   Reference[401].Actionpoint_2[7] := '0';
   Reference[401].Actionpoint_2[6] := '0';
   Reference[401].Actionpoint_2[5] := '0';
   Reference[401].Actionpoint_2[4] := '0';
   Reference[401].Actionpoint_2[3] := '0';
   Reference[401].Actionpoint_2[2] := '0';
   Reference[401].Actionpoint_2[1] := '0';
   Reference[401].Actionpoint_1[16] := '0';
   Reference[401].Actionpoint_1[15] := '0';
   Reference[401].Actionpoint_1[14] := '0';
   Reference[401].Actionpoint_1[13] := '0';
   Reference[401].Actionpoint_1[12] := '0';
   Reference[401].Actionpoint_1[11] := '0';
   Reference[401].Actionpoint_1[10] := '0';
   Reference[401].Actionpoint_1[9] := '0';
   Reference[401].Actionpoint_1[8] := '0';
   Reference[401].Actionpoint_1[7] := '0';
   Reference[401].Actionpoint_1[6] := '0';
   Reference[401].Actionpoint_1[5] := '0';
   Reference[401].Actionpoint_1[4] := '0';
   Reference[401].Actionpoint_1[3] := '0';
   Reference[401].Actionpoint_1[2] := '0';
   Reference[401].Actionpoint_1[1] := '0';
   Reference[401].Sektion[1] := 'b';
   Reference[401].Sektion[2] := 'u';
   Reference[401].Sektion[3] := 'f';
   Reference[401].Sektion[4] := 'f';
   Reference[401].Sektion[5] := 'e';
   Reference[401].Sektion[6] := 'r';
   Reference[401].Sektion[7] := '$00';
   Reference[401].Sektion[8] := '$00';
   Reference[401].Sektion[9] := '$00';
   Reference[401].Sektion[10] := '$00';
   Reference[401].Sektion[11] := '$00';
   Reference[401].Sektion[12] := '$00';
   Reference[401].Sektion[13] := '$00';
   Reference[401].Sektion[14] := '$00';
   Reference[401].Sektion[15] := '$00';
   Reference[401].Sektion[16] := '$00';
   // 19800 more start values not shown
END_DATA_BLOCK

DATA_BLOCK "DB_SDC_TS_REFERENCE_6"   // DB3785
{ S7_Optimized_Access := 'FALSE' }
VERSION : 0.1
   VAR
      HEADER : Struct   // Struktur für Datenheader // nicht verschieben
         DB_NR : Int := 3785;   // DB Nummer
         MIN_NR_SEK : Int := 501;   // Niedrigste SEK Nummer im DB
         MAX_NR_SEK : Int := 600;   // Höchste SEK Nummer im DB
         START_DAT : Int := 20;   // Startadresse der SEK im DB
         LAENGE_SEK_DATA : Int := 200;   // Länge SEK Data
         Res10 : Int := 0;   // Reserve
         Res12 : Int := 0;   // Reserve
         Res14 : Int := 0;   // Reserve
         Res16 : Int := 0;   // Reserve
         Res18 : Int := 0;   // Reserve
      END_STRUCT;
      Reference : Array[501..600] of Struct   // Sektionsnummer
         Sektion : Array[1..16] of Char;   // definition Sektion
         Actionpoint_1 : Array[1..16] of Char;   // definition Actionpoint 1
         Actionpoint_2 : Array[1..16] of Char;   // definition Actionpoint 2
         Height : Array[1..16] of Char;   // definition Hubposition (mm)
         Hoist_offset_1 : Array[1..16] of Char;   // definition Hub-Offset 1 (mm)
         Hoist_offset_2 : Array[1..16] of Char;   // definition Hub-Offset 2 (mm)
         Hoist_offset_3 : Array[1..16] of Char;   // definition Hub-Offset 3(mm)
         Hoist_offset_4 : Array[1..16] of Char;   // definition Hub-Offset 4 (mm)
         Reserve : Array[128..199] of Char;
      END_STRUCT;
   END_VAR
BEGIN
   Reference[501].Reserve[199] := ' ';
   Reference[501].Reserve[198] := ' ';
   Reference[501].Reserve[197] := ' ';
   Reference[501].Reserve[196] := ' ';
   Reference[501].Reserve[195] := ' ';
   Reference[501].Reserve[194] := ' ';
   Reference[501].Reserve[193] := ' ';
   Reference[501].Reserve[192] := ' ';
   Reference[501].Reserve[191] := ' ';
   Reference[501].Reserve[190] := ' ';
   Reference[501].Reserve[189] := ' ';
   Reference[501].Reserve[188] := ' ';
   Reference[501].Reserve[187] := ' ';
   Reference[501].Reserve[186] := ' ';
   Reference[501].Reserve[185] := ' ';
   Reference[501].Reserve[184] := ' ';
   Reference[501].Reserve[183] := ' ';
   Reference[501].Reserve[182] := ' ';
   Reference[501].Reserve[181] := ' ';
   Reference[501].Reserve[180] := ' ';
   Reference[501].Reserve[179] := ' ';
   Reference[501].Reserve[178] := ' ';
   Reference[501].Reserve[177] := ' ';
   Reference[501].Reserve[176] := ' ';
   Reference[501].Reserve[175] := ' ';
   Reference[501].Reserve[174] := ' ';
   Reference[501].Reserve[173] := ' ';
   Reference[501].Reserve[172] := ' ';
   Reference[501].Reserve[171] := ' ';
   Reference[501].Reserve[170] := ' ';
   Reference[501].Reserve[169] := ' ';
   Reference[501].Reserve[168] := ' ';
   Reference[501].Reserve[167] := ' ';
   Reference[501].Reserve[166] := ' ';
   Reference[501].Reserve[165] := ' ';
   Reference[501].Reserve[164] := ' ';
   Reference[501].Reserve[163] := ' ';
   Reference[501].Reserve[162] := ' ';
   Reference[501].Reserve[161] := ' ';
   Reference[501].Reserve[160] := ' ';
   Reference[501].Reserve[159] := ' ';
   Reference[501].Reserve[158] := ' ';
   Reference[501].Reserve[157] := ' ';
   Reference[501].Reserve[156] := ' ';
   Reference[501].Reserve[155] := ' ';
   Reference[501].Reserve[154] := ' ';
   Reference[501].Reserve[153] := ' ';
   Reference[501].Reserve[152] := ' ';
   Reference[501].Reserve[151] := ' ';
   Reference[501].Reserve[150] := ' ';
   Reference[501].Reserve[149] := ' ';
   Reference[501].Reserve[148] := ' ';
   Reference[501].Reserve[147] := ' ';
   Reference[501].Reserve[146] := ' ';
   Reference[501].Reserve[145] := ' ';
   Reference[501].Reserve[144] := ' ';
   Reference[501].Reserve[143] := '0';
   Reference[501].Reserve[142] := '0';
   Reference[501].Reserve[141] := '0';
   Reference[501].Reserve[140] := '0';
   Reference[501].Reserve[139] := '0';
   Reference[501].Reserve[138] := '0';
   Reference[501].Reserve[137] := '0';
   Reference[501].Reserve[136] := '0';
   Reference[501].Reserve[135] := '0';
   Reference[501].Reserve[134] := '0';
   Reference[501].Reserve[133] := '0';
   Reference[501].Reserve[132] := '0';
   Reference[501].Reserve[131] := '0';
   Reference[501].Reserve[130] := '0';
   Reference[501].Reserve[129] := '0';
   Reference[501].Reserve[128] := '0';
   Reference[501].Hoist_offset_4[16] := '$00';
   Reference[501].Hoist_offset_4[15] := '$00';
   Reference[501].Hoist_offset_4[14] := '$00';
   Reference[501].Hoist_offset_4[13] := '$00';
   Reference[501].Hoist_offset_4[12] := '$00';
   Reference[501].Hoist_offset_4[11] := '$00';
   Reference[501].Hoist_offset_4[10] := '$00';
   Reference[501].Hoist_offset_4[9] := '$00';
   Reference[501].Hoist_offset_4[8] := '$00';
   Reference[501].Hoist_offset_4[7] := '$00';
   Reference[501].Hoist_offset_4[6] := '$00';
   Reference[501].Hoist_offset_4[5] := '$00';
   Reference[501].Hoist_offset_4[4] := '$00';
   Reference[501].Hoist_offset_4[3] := '$00';
   Reference[501].Hoist_offset_4[2] := '$00';
   Reference[501].Hoist_offset_4[1] := '$00';
   Reference[501].Hoist_offset_3[16] := '$00';
   Reference[501].Hoist_offset_3[15] := '$00';
   Reference[501].Hoist_offset_3[14] := '$00';
   Reference[501].Hoist_offset_3[13] := '$00';
   Reference[501].Hoist_offset_3[12] := '$00';
   Reference[501].Hoist_offset_3[11] := '$00';
   Reference[501].Hoist_offset_3[10] := '$00';
   Reference[501].Hoist_offset_3[9] := '$00';
   Reference[501].Hoist_offset_3[8] := '$00';
   Reference[501].Hoist_offset_3[7] := '$00';
   Reference[501].Hoist_offset_3[6] := '$00';
   Reference[501].Hoist_offset_3[5] := '$00';
   Reference[501].Hoist_offset_3[4] := '$00';
   Reference[501].Hoist_offset_3[3] := '$00';
   Reference[501].Hoist_offset_3[2] := '$00';
   Reference[501].Hoist_offset_3[1] := '$00';
   Reference[501].Hoist_offset_2[16] := '$00';
   Reference[501].Hoist_offset_2[15] := '$00';
   Reference[501].Hoist_offset_2[14] := '$00';
   Reference[501].Hoist_offset_2[13] := '$00';
   Reference[501].Hoist_offset_2[12] := '$00';
   Reference[501].Hoist_offset_2[11] := '$00';
   Reference[501].Hoist_offset_2[10] := '$00';
   Reference[501].Hoist_offset_2[9] := '$00';
   Reference[501].Hoist_offset_2[8] := '$00';
   Reference[501].Hoist_offset_2[7] := '$00';
   Reference[501].Hoist_offset_2[6] := '$00';
   Reference[501].Hoist_offset_2[5] := '$00';
   Reference[501].Hoist_offset_2[4] := '$00';
   Reference[501].Hoist_offset_2[3] := '$00';
   Reference[501].Hoist_offset_2[2] := '$00';
   Reference[501].Hoist_offset_2[1] := '$00';
   Reference[501].Hoist_offset_1[16] := '$00';
   Reference[501].Hoist_offset_1[15] := '$00';
   Reference[501].Hoist_offset_1[14] := '$00';
   Reference[501].Hoist_offset_1[13] := '$00';
   Reference[501].Hoist_offset_1[12] := '$00';
   Reference[501].Hoist_offset_1[11] := '$00';
   Reference[501].Hoist_offset_1[10] := '$00';
   Reference[501].Hoist_offset_1[9] := '$00';
   Reference[501].Hoist_offset_1[8] := '$00';
   Reference[501].Hoist_offset_1[7] := '$00';
   Reference[501].Hoist_offset_1[6] := '$00';
   Reference[501].Hoist_offset_1[5] := '$00';
   Reference[501].Hoist_offset_1[4] := '$00';
   Reference[501].Hoist_offset_1[3] := '$00';
   Reference[501].Hoist_offset_1[2] := '$00';
   Reference[501].Hoist_offset_1[1] := '$00';
   Reference[501].Height[16] := '$00';
   Reference[501].Height[15] := '$00';
   Reference[501].Height[14] := '$00';
   Reference[501].Height[13] := '$00';
   Reference[501].Height[12] := '$00';
   Reference[501].Height[11] := '$00';
   Reference[501].Height[10] := '$00';
   Reference[501].Height[9] := '$00';
   Reference[501].Height[8] := '$00';
   Reference[501].Height[7] := '$00';
   Reference[501].Height[6] := '$00';
   Reference[501].Height[5] := '$00';
   Reference[501].Height[4] := '$00';
   Reference[501].Height[3] := '$00';
   Reference[501].Height[2] := '$00';
   Reference[501].Height[1] := '$00';
   Reference[501].Actionpoint_2[16] := '0';
   Reference[501].Actionpoint_2[15] := '0';
   Reference[501].Actionpoint_2[14] := '0';
   Reference[501].Actionpoint_2[13] := '0';
   Reference[501].Actionpoint_2[12] := '0';
   Reference[501].Actionpoint_2[11] := '0';
   Reference[501].Actionpoint_2[10] := '0';
   Reference[501].Actionpoint_2[9] := '0';
   Reference[501].Actionpoint_2[8] := '0';
   Reference[501].Actionpoint_2[7] := '0';
   Reference[501].Actionpoint_2[6] := '0';
   Reference[501].Actionpoint_2[5] := '0';
   Reference[501].Actionpoint_2[4] := '0';
   Reference[501].Actionpoint_2[3] := '0';
   Reference[501].Actionpoint_2[2] := '0';
   Reference[501].Actionpoint_2[1] := '0';
   Reference[501].Actionpoint_1[16] := '0';
   Reference[501].Actionpoint_1[15] := '0';
   Reference[501].Actionpoint_1[14] := '0';
   Reference[501].Actionpoint_1[13] := '0';
   Reference[501].Actionpoint_1[12] := '0';
   Reference[501].Actionpoint_1[11] := '0';
   Reference[501].Actionpoint_1[10] := '0';
   Reference[501].Actionpoint_1[9] := '0';
   Reference[501].Actionpoint_1[8] := '0';
   Reference[501].Actionpoint_1[7] := '0';
   Reference[501].Actionpoint_1[6] := '0';
   Reference[501].Actionpoint_1[5] := '0';
   Reference[501].Actionpoint_1[4] := '0';
   Reference[501].Actionpoint_1[3] := '0';
   Reference[501].Actionpoint_1[2] := '0';
   Reference[501].Actionpoint_1[1] := '0';
   Reference[501].Sektion[1] := 'b';
   Reference[501].Sektion[2] := 'u';
   Reference[501].Sektion[3] := 'f';
   Reference[501].Sektion[4] := 'f';
   Reference[501].Sektion[5] := 'e';
   Reference[501].Sektion[6] := 'r';
   Reference[501].Sektion[7] := '$00';
   Reference[501].Sektion[8] := '$00';
   Reference[501].Sektion[9] := '$00';
   Reference[501].Sektion[10] := '$00';
   Reference[501].Sektion[11] := '$00';
   Reference[501].Sektion[12] := '$00';
   Reference[501].Sektion[13] := '$00';
   Reference[501].Sektion[14] := '$00';
   Reference[501].Sektion[15] := '$00';
   Reference[501].Sektion[16] := '$00';
   // 19800 more start values not shown
END_DATA_BLOCK

DATA_BLOCK "DB_SDC_GLOBAL_REFERENCE"   // DB3786
{ S7_Optimized_Access := 'FALSE' }
VERSION : 0.1
   VAR
      HEADER : Struct   // Struktur für Datenheader // nicht verschieben
         DB_NR : Int := 3786;   // DB Nummer
         MIN_PAR_SET : Int := 1;   // Niedrigste PAR_SET im DB
         MAX_PAR_SET : Int := 16;   // Höchste PAR_SET im DB
         START_PAR_SET : Int := 20;   // Startadresse PAR_SET im DB
         LAENGE_PAR_SET : Int := 32;   // Länge PAR_SET im DB
         MIN_PROFIL : Int := 1;   // Niedrigste PROFIL im DB
         MAX_PROFIL : Int := 10;   // Höchste PROFIL im DB
         START_PROFIL : Int := 532;   // Startadresse PAR_SET im DB
         LAENGE_PROFIL : Int := 6;   // Länge PAR_SET im DB
         Res18 : Int := 0;   // Reserve
      END_STRUCT;
      PAR_SET : Array[0..15] of Struct
         SYNCH : Array[1..16] of Char;
         LIMITS : Array[1..16] of Char;
      END_STRUCT;
      PROFIL : Array[1..10] of Struct
         SORTE : Array[1..6] of Char;
      END_STRUCT;
   END_VAR
BEGIN
   PAR_SET[0].SYNCH[1] := 'P';
   PAR_SET[0].SYNCH[2] := 'u';
   PAR_SET[0].SYNCH[3] := 'f';
   PAR_SET[0].SYNCH[4] := 'f';
   PAR_SET[0].SYNCH[5] := 'e';
   PAR_SET[0].SYNCH[6] := 'r';
   PAR_SET[0].SYNCH[7] := 'b';
   PAR_SET[0].SYNCH[9] := 'r';
   PAR_SET[0].SYNCH[10] := 'e';
   PAR_SET[0].SYNCH[11] := 'i';
   PAR_SET[0].SYNCH[12] := 'c';
   PAR_SET[0].SYNCH[13] := 'h';
   PAR_SET[0].SYNCH[14] := '$00';
   PAR_SET[0].SYNCH[15] := '$00';
   PAR_SET[0].SYNCH[16] := '$00';
   PAR_SET[1].SYNCH[1] := 'A';
   PAR_SET[1].SYNCH[2] := 'r';
   PAR_SET[1].SYNCH[3] := 'b';
   PAR_SET[1].SYNCH[4] := 'e';
   PAR_SET[1].SYNCH[5] := 'i';
   PAR_SET[1].SYNCH[6] := 's';
   PAR_SET[1].SYNCH[7] := 't';
   PAR_SET[1].SYNCH[8] := 'l';
   PAR_SET[1].SYNCH[9] := 'i';
   PAR_SET[1].SYNCH[10] := 'n';
   PAR_SET[1].SYNCH[11] := 'i';
   PAR_SET[1].SYNCH[12] := 'e';
   PAR_SET[1].SYNCH[13] := '$00';
   PAR_SET[1].SYNCH[14] := '$00';
   PAR_SET[1].SYNCH[15] := '$00';
   PAR_SET[1].SYNCH[16] := '$00';
   PAR_SET[2].SYNCH[1] := 'A';
   PAR_SET[2].SYNCH[2] := 'n';
   PAR_SET[2].SYNCH[3] := 'd';
   PAR_SET[2].SYNCH[4] := 'o';
   PAR_SET[2].SYNCH[5] := 'c';
   PAR_SET[2].SYNCH[6] := 'k';
   PAR_SET[2].SYNCH[8] := 'e';
   PAR_SET[2].SYNCH[9] := 'r';
   PAR_SET[2].SYNCH[10] := 'e';
   PAR_SET[2].SYNCH[11] := 'i';
   PAR_SET[2].SYNCH[12] := 'c';
   PAR_SET[2].SYNCH[13] := 'h';
   PAR_SET[2].SYNCH[14] := '$00';
   PAR_SET[2].SYNCH[15] := '$00';
   PAR_SET[2].SYNCH[16] := '$00';
   PAR_SET[3].SYNCH[1] := 'A';
   PAR_SET[3].SYNCH[2] := 'b';
   PAR_SET[3].SYNCH[3] := 'z';
   PAR_SET[3].SYNCH[4] := 'u';
   PAR_SET[3].SYNCH[5] := 'g';
   PAR_SET[3].SYNCH[6] := 's';
   PAR_SET[3].SYNCH[7] := 'b';
   PAR_SET[3].SYNCH[8] := 'e';
   PAR_SET[3].SYNCH[9] := 'r';
   PAR_SET[3].SYNCH[10] := 'e';
   PAR_SET[3].SYNCH[11] := 'i';
   PAR_SET[3].SYNCH[12] := 'c';
   PAR_SET[3].SYNCH[13] := 'h';
   PAR_SET[3].SYNCH[14] := '$00';
   PAR_SET[3].SYNCH[15] := '$00';
   PAR_SET[3].SYNCH[16] := '$00';
   PAR_SET[4].SYNCH[1] := 'A';
   PAR_SET[4].SYNCH[2] := 'n';
   PAR_SET[4].SYNCH[3] := 'd';
   PAR_SET[4].SYNCH[4] := '.';
   PAR_SET[4].SYNCH[5] := ' ';
   PAR_SET[4].SYNCH[6] := 'A';
   PAR_SET[4].SYNCH[7] := 'r';
   PAR_SET[4].SYNCH[8] := 'b';
   PAR_SET[4].SYNCH[9] := 'e';
   PAR_SET[4].SYNCH[10] := 'i';
   PAR_SET[4].SYNCH[11] := 't';
   PAR_SET[4].SYNCH[12] := 's';
   PAR_SET[4].SYNCH[13] := 'p';
   PAR_SET[4].SYNCH[14] := 'l';
   PAR_SET[4].SYNCH[15] := 'a';
   PAR_SET[4].SYNCH[16] := 't';
   PAR_SET[5].SYNCH[1] := 'K';
   PAR_SET[5].SYNCH[2] := 'u';
   PAR_SET[5].SYNCH[3] := 'r';
   PAR_SET[5].SYNCH[4] := 'v';
   PAR_SET[5].SYNCH[5] := 'e';
   PAR_SET[5].SYNCH[6] := '$00';
   PAR_SET[5].SYNCH[7] := '$00';
   PAR_SET[5].SYNCH[8] := '$00';
   PAR_SET[5].SYNCH[9] := '$00';
   PAR_SET[5].SYNCH[10] := '$00';
   PAR_SET[5].SYNCH[11] := '$00';
   PAR_SET[5].SYNCH[12] := '$00';
   PAR_SET[5].SYNCH[13] := '$00';
   PAR_SET[5].SYNCH[14] := '$00';
   PAR_SET[5].SYNCH[15] := '$00';
   PAR_SET[5].SYNCH[16] := '$00';
   PAR_SET[6].SYNCH[1] := 'v';
   PAR_SET[6].SYNCH[2] := 'o';
   PAR_SET[6].SYNCH[3] := 'r';
   PAR_SET[6].SYNCH[4] := ' ';
   PAR_SET[6].SYNCH[5] := 'K';
   PAR_SET[6].SYNCH[6] := 'u';
   PAR_SET[6].SYNCH[7] := 'r';
   PAR_SET[6].SYNCH[8] := 'v';
   PAR_SET[6].SYNCH[9] := 'e';
   PAR_SET[6].SYNCH[10] := '$00';
   PAR_SET[6].SYNCH[11] := '$00';
   PAR_SET[6].SYNCH[12] := '$00';
   PAR_SET[6].SYNCH[13] := '$00';
   PAR_SET[6].SYNCH[14] := '$00';
   PAR_SET[6].SYNCH[15] := '$00';
   PAR_SET[6].SYNCH[16] := '$00';
   PAR_SET[7].SYNCH[1] := 'n';
   PAR_SET[7].SYNCH[2] := 'a';
   PAR_SET[7].SYNCH[3] := 'c';
   PAR_SET[7].SYNCH[4] := 'h';
   PAR_SET[7].SYNCH[5] := ' ';
   PAR_SET[7].SYNCH[6] := 'K';
   PAR_SET[7].SYNCH[7] := 'u';
   PAR_SET[7].SYNCH[8] := 'r';
   PAR_SET[7].SYNCH[9] := 'v';
   PAR_SET[7].SYNCH[10] := 'e';
   PAR_SET[7].SYNCH[11] := '$00';
   PAR_SET[7].SYNCH[12] := '$00';
   PAR_SET[7].SYNCH[13] := '$00';
   PAR_SET[7].SYNCH[14] := '$00';
   PAR_SET[7].SYNCH[15] := '$00';
   PAR_SET[7].SYNCH[16] := '$00';
   PAR_SET[8].SYNCH[1] := 'R';
   PAR_SET[8].SYNCH[2] := 'e';
   PAR_SET[8].SYNCH[3] := 's';
   PAR_SET[8].SYNCH[4] := 'e';
   PAR_SET[8].SYNCH[5] := 'r';
   PAR_SET[8].SYNCH[6] := 'v';
   PAR_SET[8].SYNCH[7] := 'e';
   PAR_SET[8].SYNCH[8] := '$00';
   PAR_SET[8].SYNCH[9] := '$00';
   PAR_SET[8].SYNCH[10] := '$00';
   PAR_SET[8].SYNCH[11] := '$00';
   PAR_SET[8].SYNCH[12] := '$00';
   PAR_SET[8].SYNCH[13] := '$00';
   PAR_SET[8].SYNCH[14] := '$00';
   PAR_SET[8].SYNCH[15] := '$00';
   PAR_SET[8].SYNCH[16] := '$00';
   PAR_SET[9].SYNCH[1] := 'H';
   PAR_SET[9].SYNCH[2] := 'e';
   PAR_SET[9].SYNCH[3] := 'b';
   PAR_SET[9].SYNCH[4] := 'e';
   PAR_SET[9].SYNCH[5] := 'r';
   PAR_SET[9].SYNCH[6] := '$00';
   PAR_SET[9].SYNCH[7] := '$00';
   PAR_SET[9].SYNCH[8] := '$00';
   PAR_SET[9].SYNCH[9] := '$00';
   PAR_SET[9].SYNCH[10] := '$00';
   PAR_SET[9].SYNCH[11] := '$00';
   PAR_SET[9].SYNCH[12] := '$00';
   PAR_SET[9].SYNCH[13] := '$00';
   PAR_SET[9].SYNCH[14] := '$00';
   PAR_SET[9].SYNCH[15] := '$00';
   PAR_SET[9].SYNCH[16] := '$00';
   PAR_SET[10].SYNCH[1] := 'T';
   PAR_SET[10].SYNCH[2] := 'e';
   PAR_SET[10].SYNCH[3] := 'c';
   PAR_SET[10].SYNCH[4] := 'h';
   PAR_SET[10].SYNCH[5] := 'n';
   PAR_SET[10].SYNCH[6] := 'i';
   PAR_SET[10].SYNCH[7] := 'k';
   PAR_SET[10].SYNCH[8] := 't';
   PAR_SET[10].SYNCH[9] := 'a';
   PAR_SET[10].SYNCH[10] := 'c';
   PAR_SET[10].SYNCH[11] := 'k';
   PAR_SET[10].SYNCH[12] := 't';
   PAR_SET[10].SYNCH[13] := '$00';
   PAR_SET[10].SYNCH[14] := '$00';
   PAR_SET[10].SYNCH[15] := '$00';
   PAR_SET[10].SYNCH[16] := '$00';
   PAR_SET[11].SYNCH[1] := 'K';
   PAR_SET[11].SYNCH[2] := 'u';
   PAR_SET[11].SYNCH[3] := 'r';
   PAR_SET[11].SYNCH[4] := 'v';
   PAR_SET[11].SYNCH[5] := 'e';
   PAR_SET[11].SYNCH[6] := ' ';
   PAR_SET[11].SYNCH[7] := 'l';
   PAR_SET[11].SYNCH[8] := 'e';
   PAR_SET[11].SYNCH[9] := 'e';
   PAR_SET[11].SYNCH[10] := 'r';
   PAR_SET[11].SYNCH[11] := '$00';
   PAR_SET[11].SYNCH[12] := '$00';
   PAR_SET[11].SYNCH[13] := '$00';
   PAR_SET[11].SYNCH[14] := '$00';
   PAR_SET[11].SYNCH[15] := '$00';
   PAR_SET[11].SYNCH[16] := '$00';
   PAR_SET[12].SYNCH[1] := 'F';
   PAR_SET[12].SYNCH[2] := 'r';
   PAR_SET[12].SYNCH[3] := 'o';
   PAR_SET[12].SYNCH[4] := 'n';
   PAR_SET[12].SYNCH[5] := 't';
   PAR_SET[12].SYNCH[6] := 'e';
   PAR_SET[12].SYNCH[7] := 'n';
   PAR_SET[12].SYNCH[8] := 'd';
   PAR_SET[12].SYNCH[9] := ' ';
   PAR_SET[12].SYNCH[10] := 'A';
   // 372 more start values not shown
END_DATA_BLOCK

DATA_BLOCK "DB_SDC_EMS_FLAGS_HMI"   // DB3801
{ S7_Optimized_Access := 'FALSE' }
AUTHOR : FFM
FAMILY : SDC
NAME : GLOBAL
VERSION : 0.1
   VAR
      HEADER : Struct
         DB_NR : Int := 3801;
         Res020 : Int := 0;
         Res040 : Int := 0;
         START_EMS : Int := 20;
         LAENGE_EMS_FLAGS : Int := 2;
         START_HMI : Int := 20;
         OFFEST_HMI_DATA : Int := 20;
         Res140 : Int := 0;
         Res160 : Int := 0;
         Res180 : Int := 0;
      END_STRUCT;
      HMI : Array[1..30] of Struct
         PULT_Nr_EDIT : Int;
         BILD_Nr : Int;
         BILD_Nr_Alt : Int;
         EMS_Nr : Int;
         EMS_Nr_Alt : Int;
         TIME_SFC12 : Int;
         LADDR_SFC12 : Hw_Any;
         RET_VAL_SFC12 : Int;
         MODE_SFC12 : Byte;
         RES17 : Byte;
         T_EDIT : Bool;
         T_RESET_BED : Bool;
         T_SAVE : Bool;
         T_LOAD : Bool;
         T_ACTIV : Bool;
         T_DEACTIV : Bool;
         Res086 : Bool;
         Res087 : Bool;
         FR_EDIT : Bool;
         ER_DATA : Bool;
         BUSY_SFC12 : Bool;
         REQ_SFC12 : Bool;
         FLAGS : "UDT_SDC_EMS_FLAGS";
      END_STRUCT;
   END_VAR
BEGIN
   HMI[1].PULT_Nr_EDIT := 0;
   HMI[1].BILD_Nr := 0;
   HMI[1].BILD_Nr_Alt := 0;
   HMI[1].EMS_Nr := 1;
   HMI[1].EMS_Nr_Alt := 0;
   HMI[1].TIME_SFC12 := 31;
   HMI[1].LADDR_SFC12 := 16#01C9;
   HMI[1].RET_VAL_SFC12 := 28672;
   HMI[1].MODE_SFC12 := 16#01;
   HMI[1].RES17 := 16#00;
   HMI[1].T_EDIT := FALSE;
   HMI[1].T_RESET_BED := FALSE;
   HMI[1].T_SAVE := FALSE;
   HMI[1].T_LOAD := FALSE;
   HMI[1].T_ACTIV := FALSE;
   HMI[1].T_DEACTIV := FALSE;
   HMI[1].Res086 := FALSE;
   HMI[1].Res087 := FALSE;
   HMI[1].FR_EDIT := FALSE;
   HMI[1].ER_DATA := FALSE;
   HMI[1].BUSY_SFC12 := FALSE;
   HMI[1].REQ_SFC12 := FALSE;
   HMI[1].FLAGS.PRESENT := FALSE;
   HMI[1].FLAGS.IN_HW := FALSE;
   HMI[1].FLAGS.ACTIV := FALSE;
   HMI[1].FLAGS.ENABLE := FALSE;
   HMI[1].FLAGS.COMM_FAULT := FALSE;
   HMI[1].FLAGS.FAULTY := FALSE;
   HMI[1].FLAGS.SIMULATION := FALSE;
   HMI[1].FLAGS.Spare_0_7 := FALSE;
   HMI[1].FLAGS.Spare_1_0 := FALSE;
   HMI[1].FLAGS.Spare_1_1 := FALSE;
   HMI[1].FLAGS.Spare_1_2 := FALSE;
   HMI[1].FLAGS.Spare_1_3 := FALSE;
   HMI[1].FLAGS.Spare_1_4 := FALSE;
   HMI[1].FLAGS.Spare_1_5 := FALSE;
   HMI[1].FLAGS.Spare_1_6 := FALSE;
   HMI[1].FLAGS.Spare_1_7 := FALSE;
   HMI[2].PULT_Nr_EDIT := 0;
   HMI[2].BILD_Nr := 0;
   HMI[2].BILD_Nr_Alt := 0;
   HMI[2].EMS_Nr := 1;
   HMI[2].EMS_Nr_Alt := 1;
   HMI[2].TIME_SFC12 := 0;
   HMI[2].LADDR_SFC12 := 16#0000;
   HMI[2].RET_VAL_SFC12 := 0;
   HMI[2].MODE_SFC12 := 16#00;
   HMI[2].RES17 := 16#00;
   HMI[2].T_EDIT := FALSE;
   HMI[2].T_RESET_BED := FALSE;
   HMI[2].T_SAVE := FALSE;
   HMI[2].T_LOAD := FALSE;
   HMI[2].T_ACTIV := FALSE;
   HMI[2].T_DEACTIV := FALSE;
   HMI[2].Res086 := FALSE;
   HMI[2].Res087 := FALSE;
   HMI[2].FR_EDIT := FALSE;
   HMI[2].ER_DATA := FALSE;
   HMI[2].BUSY_SFC12 := FALSE;
   HMI[2].REQ_SFC12 := FALSE;
   HMI[2].FLAGS.PRESENT := TRUE;
   HMI[2].FLAGS.IN_HW := TRUE;
   HMI[2].FLAGS.ACTIV := TRUE;
   HMI[2].FLAGS.ENABLE := FALSE;
   HMI[2].FLAGS.COMM_FAULT := FALSE;
   HMI[2].FLAGS.FAULTY := TRUE;
   HMI[2].FLAGS.SIMULATION := FALSE;
   HMI[2].FLAGS.Spare_0_7 := FALSE;
   HMI[2].FLAGS.Spare_1_0 := FALSE;
   HMI[2].FLAGS.Spare_1_1 := FALSE;
   HMI[2].FLAGS.Spare_1_2 := FALSE;
   HMI[2].FLAGS.Spare_1_3 := FALSE;
   HMI[2].FLAGS.Spare_1_4 := FALSE;
   HMI[2].FLAGS.Spare_1_5 := FALSE;
   HMI[2].FLAGS.Spare_1_6 := FALSE;
   HMI[2].FLAGS.Spare_1_7 := FALSE;
   HMI[3].PULT_Nr_EDIT := 0;
   HMI[3].BILD_Nr := 0;
   HMI[3].BILD_Nr_Alt := 0;
   HMI[3].EMS_Nr := 1;
   HMI[3].EMS_Nr_Alt := 0;
   HMI[3].TIME_SFC12 := 0;
   HMI[3].LADDR_SFC12 := 16#0000;
   HMI[3].RET_VAL_SFC12 := 0;
   HMI[3].MODE_SFC12 := 16#00;
   HMI[3].RES17 := 16#00;
   HMI[3].T_EDIT := FALSE;
   HMI[3].T_RESET_BED := FALSE;
   HMI[3].T_SAVE := FALSE;
   HMI[3].T_LOAD := FALSE;
   HMI[3].T_ACTIV := FALSE;
   HMI[3].T_DEACTIV := FALSE;
   HMI[3].Res086 := FALSE;
   HMI[3].Res087 := FALSE;
   HMI[3].FR_EDIT := FALSE;
   HMI[3].ER_DATA := FALSE;
   HMI[3].BUSY_SFC12 := FALSE;
   HMI[3].REQ_SFC12 := FALSE;
   HMI[3].FLAGS.PRESENT := FALSE;
   HMI[3].FLAGS.IN_HW := FALSE;
   HMI[3].FLAGS.ACTIV := FALSE;
   HMI[3].FLAGS.ENABLE := FALSE;
   HMI[3].FLAGS.COMM_FAULT := FALSE;
   HMI[3].FLAGS.FAULTY := FALSE;
   HMI[3].FLAGS.SIMULATION := FALSE;
   HMI[3].FLAGS.Spare_0_7 := FALSE;
   HMI[3].FLAGS.Spare_1_0 := FALSE;
   HMI[3].FLAGS.Spare_1_1 := FALSE;
   HMI[3].FLAGS.Spare_1_2 := FALSE;
   HMI[3].FLAGS.Spare_1_3 := FALSE;
   HMI[3].FLAGS.Spare_1_4 := FALSE;
   HMI[3].FLAGS.Spare_1_5 := FALSE;
   HMI[3].FLAGS.Spare_1_6 := FALSE;
   HMI[3].FLAGS.Spare_1_7 := FALSE;
   HMI[4].PULT_Nr_EDIT := 0;
   HMI[4].BILD_Nr := 0;
   HMI[4].BILD_Nr_Alt := 0;
   HMI[4].EMS_Nr := 1;
   HMI[4].EMS_Nr_Alt := 0;
   HMI[4].TIME_SFC12 := 0;
   HMI[4].LADDR_SFC12 := 16#0000;
   HMI[4].RET_VAL_SFC12 := 0;
   HMI[4].MODE_SFC12 := 16#00;
   HMI[4].RES17 := 16#00;
   HMI[4].T_EDIT := FALSE;
   HMI[4].T_RESET_BED := FALSE;
   HMI[4].T_SAVE := FALSE;
   HMI[4].T_LOAD := FALSE;
   HMI[4].T_ACTIV := FALSE;
   HMI[4].T_DEACTIV := FALSE;
   HMI[4].Res086 := FALSE;
   HMI[4].Res087 := FALSE;
   HMI[4].FR_EDIT := FALSE;
   HMI[4].ER_DATA := FALSE;
   HMI[4].BUSY_SFC12 := FALSE;
   HMI[4].REQ_SFC12 := FALSE;
   HMI[4].FLAGS.PRESENT := FALSE;
   HMI[4].FLAGS.IN_HW := FALSE;
   HMI[4].FLAGS.ACTIV := FALSE;
   HMI[4].FLAGS.ENABLE := FALSE;
   HMI[4].FLAGS.COMM_FAULT := FALSE;
   HMI[4].FLAGS.FAULTY := FALSE;
   HMI[4].FLAGS.SIMULATION := FALSE;
   HMI[4].FLAGS.Spare_0_7 := FALSE;
   HMI[4].FLAGS.Spare_1_0 := FALSE;
   HMI[4].FLAGS.Spare_1_1 := FALSE;
   HMI[4].FLAGS.Spare_1_2 := FALSE;
   HMI[4].FLAGS.Spare_1_3 := FALSE;
   HMI[4].FLAGS.Spare_1_4 := FALSE;
   HMI[4].FLAGS.Spare_1_5 := FALSE;
   HMI[4].FLAGS.Spare_1_6 := FALSE;
   HMI[4].FLAGS.Spare_1_7 := FALSE;
   HMI[5].PULT_Nr_EDIT := 0;
   HMI[5].BILD_Nr := 0;
   HMI[5].BILD_Nr_Alt := 0;
   HMI[5].EMS_Nr := 0;
   HMI[5].EMS_Nr_Alt := 0;
   HMI[5].TIME_SFC12 := 0;
   HMI[5].LADDR_SFC12 := 16#0000;
   HMI[5].RET_VAL_SFC12 := 0;
   HMI[5].MODE_SFC12 := 16#00;
   HMI[5].RES17 := 16#00;
   HMI[5].T_EDIT := FALSE;
   HMI[5].T_RESET_BED := FALSE;
   HMI[5].T_SAVE := FALSE;
   HMI[5].T_LOAD := FALSE;
   HMI[5].T_ACTIV := FALSE;
   HMI[5].T_DEACTIV := FALSE;
   HMI[5].Res086 := FALSE;
   HMI[5].Res087 := FALSE;
   HMI[5].FR_EDIT := FALSE;
   HMI[5].ER_DATA := FALSE;
   HMI[5].BUSY_SFC12 := FALSE;
   HMI[5].REQ_SFC12 := FALSE;
   HMI[5].FLAGS.PRESENT := FALSE;
   HMI[5].FLAGS.IN_HW := FALSE;
   HMI[5].FLAGS.ACTIV := FALSE;
   HMI[5].FLAGS.ENABLE := FALSE;
   HMI[5].FLAGS.COMM_FAULT := FALSE;
   HMI[5].FLAGS.FAULTY := FALSE;
   HMI[5].FLAGS.SIMULATION := FALSE;
   HMI[5].FLAGS.Spare_0_7 := FALSE;
   HMI[5].FLAGS.Spare_1_0 := FALSE;
   HMI[5].FLAGS.Spare_1_1 := FALSE;
   HMI[5].FLAGS.Spare_1_2 := FALSE;
   HMI[5].FLAGS.Spare_1_3 := FALSE;
   HMI[5].FLAGS.Spare_1_4 := FALSE;
   HMI[5].FLAGS.Spare_1_5 := FALSE;
   HMI[5].FLAGS.Spare_1_6 := FALSE;
   HMI[5].FLAGS.Spare_1_7 := FALSE;
   HMI[6].PULT_Nr_EDIT := 0;
   HMI[6].BILD_Nr := 0;
   HMI[6].BILD_Nr_Alt := 0;
   HMI[6].EMS_Nr := 1;
   HMI[6].EMS_Nr_Alt := 0;
   HMI[6].TIME_SFC12 := 0;
   HMI[6].LADDR_SFC12 := 16#0000;
   HMI[6].RET_VAL_SFC12 := 0;
   HMI[6].MODE_SFC12 := 16#00;
   HMI[6].RES17 := 16#00;
   // 560 more start values not shown
END_DATA_BLOCK

DATA_BLOCK "DB_SDC_EMS_PAR_HMI"   // DB3802
{ S7_Optimized_Access := 'FALSE' }
VERSION : 0.1
   VAR
      HEADER : Struct
         DB_NR : Int := 3802;
         Res020 : Int := 0;
         Res040 : Int := 0;
         START_PAR : Int := 20;
         LAENGE_PAR : Int := 300;
         Res100 : Int := 0;
         Res120 : Int := 0;
         Res140 : Int := 0;
         START_HMI : Int := 20;
         OFFEST_HMI_DATA : Int := 20;
      END_STRUCT;
      HMI : Array[1..20] of Struct
         PULT_Nr_EDIT : Int;
         BILD_Nr : Int;
         BILD_Nr_Alt : Int;
         Res060 : Int;
         Res080 : Int;
         Res100 : Int;
         Res120 : Int;
         Res140 : Int;
         Res160 : Int;
         T_EDIT : Bool;
         T_RESET_BED : Bool;
         T_SAVE : Bool;
         T_LOAD : Bool;
         Res084 : Bool;
         Res085 : Bool;
         Res086 : Bool;
         Res087 : Bool;
         FR_EDIT : Bool;
         ER_DATA : Bool;
         PAR : "UDT_EMS_PAR";
      END_STRUCT;
   END_VAR
BEGIN
   HMI[1].PULT_Nr_EDIT := 0;
   HMI[1].BILD_Nr := 0;
   HMI[1].BILD_Nr_Alt := 0;
   HMI[1].Res060 := 0;
   HMI[1].Res080 := 0;
   HMI[1].Res100 := 0;
   HMI[1].Res120 := 0;
   HMI[1].Res140 := 0;
   HMI[1].Res160 := 0;
   HMI[1].T_EDIT := FALSE;
   HMI[1].T_RESET_BED := FALSE;
   HMI[1].T_SAVE := FALSE;
   HMI[1].T_LOAD := FALSE;
   HMI[1].Res084 := FALSE;
   HMI[1].Res085 := FALSE;
   HMI[1].Res086 := FALSE;
   HMI[1].Res087 := FALSE;
   HMI[1].FR_EDIT := FALSE;
   HMI[1].ER_DATA := FALSE;
   HMI[1].PAR.DRIVE.Funct.Res0 := TRUE;
   HMI[1].PAR.DRIVE.Funct.IgnoreBridgeStopp := TRUE;
   HMI[1].PAR.DRIVE.Funct.DontIgnoreAPOSwhenDriving := FALSE;
   HMI[1].PAR.DRIVE.Funct.Speed0_1mm_s := FALSE;
   HMI[1].PAR.DRIVE.Funct.IR_noEMSnumber := FALSE;
   HMI[1].PAR.DRIVE.Funct.IR_noLogin := FALSE;
   HMI[1].PAR.DRIVE.Funct.Res6 := FALSE;
   HMI[1].PAR.DRIVE.Funct.Res7 := FALSE;
   HMI[1].PAR.DRIVE.Funct.Res8 := FALSE;
   HMI[1].PAR.DRIVE.Funct.Res9 := FALSE;
   HMI[1].PAR.DRIVE.Funct.Res10 := FALSE;
   HMI[1].PAR.DRIVE.Funct.Res11 := FALSE;
   HMI[1].PAR.DRIVE.Funct.Res12 := FALSE;
   HMI[1].PAR.DRIVE.Funct.Res13 := FALSE;
   HMI[1].PAR.DRIVE.Funct.Res14 := FALSE;
   HMI[1].PAR.DRIVE.Funct.Res15 := FALSE;
   HMI[1].PAR.DRIVE.V_FACT_1 := 0.00296;
   HMI[1].PAR.DRIVE.V_SETP_1 := 600;
   HMI[1].PAR.DRIVE.V_FACT_2 := 0.00266;
   HMI[1].PAR.DRIVE.V_SETP_2 := 3000;
   HMI[1].PAR.DRIVE.V_FACT_3 := 0.00246;
   HMI[1].PAR.DRIVE.V_SETP_3 := 10000;
   HMI[1].PAR.DRIVE.V_FACT_4 := 0.0024;
   HMI[1].PAR.DRIVE.V_SETP_4 := 20000;
   HMI[1].PAR.DRIVE.V_LIMIT_FACT := 0.2;
   HMI[1].PAR.DRIVE.V_FACT_5 := 0.0024;
   HMI[1].PAR.DRIVE."V_FACT_ACT_V_<600" := 0.0027;
   HMI[1].PAR.DRIVE."V_FACT_ACT_V_<1200" := 0.0027;
   HMI[1].PAR.DRIVE.V_min := 300;
   HMI[1].PAR.DRIVE.V_max_top := 40000;
   HMI[1].PAR.DRIVE.V_max_Not_top := 20000;
   HMI[1].PAR.DRIVE.V_Pos_1_Reserve := 0;
   HMI[1].PAR.DRIVE.V_Pos_2 := 10000;
   HMI[1].PAR.DRIVE.V_Pos_3_Reserve := 12000;
   HMI[1].PAR.DRIVE.V_Fixed_1 := 3000;
   HMI[1].PAR.DRIVE.V_Fixed_2 := 13000;
   HMI[1].PAR.DRIVE.V_Fixed_3_Reserve := 18000;
   HMI[1].PAR.DRIVE.V_Fixed_4_SLS_SPEED := 15000;
   HMI[1].PAR.DRIVE.V_DIV_FAST := 18000;
   HMI[1].PAR.DRIVE.DIV_POS_FAST := 40;
   HMI[1].PAR.DRIVE.DIV_POS_SLOW := 60;
   HMI[1].PAR.DRIVE.TOL_SET_POS := 2;
   HMI[1].PAR.DRIVE.TOL_RESET_POS := 20;
   HMI[1].PAR.DRIVE.Window_Pos := 2;
   HMI[1].PAR.DRIVE.Window_Overrun := 10;
   HMI[1].PAR.DRIVE.Window_Pos_2 := 800;
   HMI[1].PAR.DRIVE.Window_Movement := 10;
   HMI[1].PAR.DRIVE.Window_Distance_Reserve := 10;
   HMI[1].PAR.DRIVE.Delay_Pos := 2000;
   HMI[1].PAR.DRIVE.Reserve_118 := S5T#5M;
   HMI[1].PAR.DRIVE.Reserve_120 := S5T#2M;
   HMI[1].PAR.DRIVE.DelaySpeedContr := S5T#6S_600MS;
   HMI[1].PAR.DRIVE.TolSpeedContr := 30;
   HMI[1].PAR.DRIVE.SYNCH_MID_VALUE := 0;
   HMI[1].PAR.Reserve[1] := 16#0000;
   HMI[1].PAR.Reserve[2] := 16#0000;
   HMI[1].PAR.Reserve[3] := 16#0000;
   HMI[1].PAR.Reserve[4] := 16#0000;
   HMI[1].PAR.Reserve[5] := 16#0000;
   HMI[1].PAR.HOIST.V_Min := 0;
   HMI[1].PAR.HOIST.V_Max := 8000;
   HMI[1].PAR.HOIST.V_MaxOccLift := 6500;
   HMI[1].PAR.HOIST.V_Reserve_2 := 0;
   HMI[1].PAR.HOIST.V_Pos_1 := 800;
   HMI[1].PAR.HOIST.V_Pos_2 := 2000;
   HMI[1].PAR.HOIST.V_Fixed_1 := 2000;
   HMI[1].PAR.HOIST.V_Fixed_2 := 4000;
   HMI[1].PAR.HOIST.V_Fixed_3_START := 400;
   HMI[1].PAR.HOIST.V_Fixed_4_SLS_SPEED := 2000;
   HMI[1].PAR.HOIST.V_Fixed_5_Reserve := 2000;
   HMI[1].PAR.HOIST.V_Fixed_6_SlowSpeed := 2000;
   HMI[1].PAR.HOIST.V_FACT_Hz_UP := 0.012448;
   HMI[1].PAR.HOIST.V_FACT_Hz_DOWN := 0.012462;
   HMI[1].PAR.HOIST.H_Window_POS_V1 := 20;
   HMI[1].PAR.HOIST.H_Window_POS_V2 := 140;
   HMI[1].PAR.HOIST.H_TOL_SET_POS := 1;
   HMI[1].PAR.HOIST.H_TOL_RESET_POS := 7;
   HMI[1].PAR.HOIST.H_MIN := 4;
   HMI[1].PAR.HOIST.H_MIN_without_bypass := 122;
   HMI[1].PAR.HOIST.H_REF_OFFSET := 8;
   HMI[1].PAR.HOIST.H_REF := 4151;
   HMI[1].PAR.HOIST.H_FACT_ENC1 := 1.0;
   HMI[1].PAR.HOIST.H_FACT_ENC2 := 1.0;
   HMI[1].PAR.HOIST.H_FACT_SPEED := 0.316;
   HMI[1].PAR.HOIST.H_ENC_MAX_DIFF := 50;
   HMI[1].PAR.HOIST.H_Slow := 560;
   HMI[1].PAR.HOIST.H_tIN_POS := 1000;
   HMI[1].PAR.HOIST.H_REF_HMI := 4151;
   HMI[1].PAR.Reserve1[1] := 16#0000;
   HMI[1].PAR.Reserve1[2] := 16#0000;
   HMI[1].PAR.Reserve1[3] := 16#0000;
   HMI[1].PAR.Reserve1[4] := 16#0000;
   HMI[1].PAR.Reserve1[5] := 16#0000;
   HMI[1].PAR.Reserve1[6] := 16#0000;
   HMI[2].PULT_Nr_EDIT := 0;
   HMI[2].BILD_Nr := 0;
   HMI[2].BILD_Nr_Alt := 0;
   HMI[2].Res060 := 0;
   HMI[2].Res080 := 0;
   HMI[2].Res100 := 0;
   HMI[2].Res120 := 0;
   HMI[2].Res140 := 0;
   HMI[2].Res160 := 0;
   HMI[2].T_EDIT := FALSE;
   HMI[2].T_RESET_BED := FALSE;
   HMI[2].T_SAVE := FALSE;
   HMI[2].T_LOAD := FALSE;
   HMI[2].Res084 := FALSE;
   HMI[2].Res085 := FALSE;
   HMI[2].Res086 := FALSE;
   HMI[2].Res087 := FALSE;
   HMI[2].FR_EDIT := FALSE;
   HMI[2].ER_DATA := FALSE;
   HMI[2].PAR.DRIVE.Funct.Res0 := TRUE;
   HMI[2].PAR.DRIVE.Funct.IgnoreBridgeStopp := TRUE;
   HMI[2].PAR.DRIVE.Funct.DontIgnoreAPOSwhenDriving := FALSE;
   HMI[2].PAR.DRIVE.Funct.Speed0_1mm_s := FALSE;
   HMI[2].PAR.DRIVE.Funct.IR_noEMSnumber := FALSE;
   HMI[2].PAR.DRIVE.Funct.IR_noLogin := FALSE;
   HMI[2].PAR.DRIVE.Funct.Res6 := FALSE;
   HMI[2].PAR.DRIVE.Funct.Res7 := FALSE;
   HMI[2].PAR.DRIVE.Funct.Res8 := FALSE;
   HMI[2].PAR.DRIVE.Funct.Res9 := FALSE;
   HMI[2].PAR.DRIVE.Funct.Res10 := FALSE;
   HMI[2].PAR.DRIVE.Funct.Res11 := FALSE;
   HMI[2].PAR.DRIVE.Funct.Res12 := FALSE;
   HMI[2].PAR.DRIVE.Funct.Res13 := FALSE;
   HMI[2].PAR.DRIVE.Funct.Res14 := FALSE;
   HMI[2].PAR.DRIVE.Funct.Res15 := FALSE;
   HMI[2].PAR.DRIVE.V_FACT_1 := 0.00296;
   HMI[2].PAR.DRIVE.V_SETP_1 := 600;
   HMI[2].PAR.DRIVE.V_FACT_2 := 0.00266;
   HMI[2].PAR.DRIVE.V_SETP_2 := 3000;
   HMI[2].PAR.DRIVE.V_FACT_3 := 0.00246;
   HMI[2].PAR.DRIVE.V_SETP_3 := 10000;
   HMI[2].PAR.DRIVE.V_FACT_4 := 0.0024;
   HMI[2].PAR.DRIVE.V_SETP_4 := 20000;
   HMI[2].PAR.DRIVE.V_LIMIT_FACT := 0.2;
   HMI[2].PAR.DRIVE.V_FACT_5 := 0.0024;
   HMI[2].PAR.DRIVE."V_FACT_ACT_V_<600" := 0.0027;
   HMI[2].PAR.DRIVE."V_FACT_ACT_V_<1200" := 0.0027;
   HMI[2].PAR.DRIVE.V_min := 300;
   HMI[2].PAR.DRIVE.V_max_top := 40000;
   HMI[2].PAR.DRIVE.V_max_Not_top := 20000;
   HMI[2].PAR.DRIVE.V_Pos_1_Reserve := 0;
   HMI[2].PAR.DRIVE.V_Pos_2 := 10000;
   HMI[2].PAR.DRIVE.V_Pos_3_Reserve := 12000;
   HMI[2].PAR.DRIVE.V_Fixed_1 := 3000;
   HMI[2].PAR.DRIVE.V_Fixed_2 := 13000;
   HMI[2].PAR.DRIVE.V_Fixed_3_Reserve := 18000;
   HMI[2].PAR.DRIVE.V_Fixed_4_SLS_SPEED := 15000;
   HMI[2].PAR.DRIVE.V_DIV_FAST := 18000;
   HMI[2].PAR.DRIVE.DIV_POS_FAST := 40;
   HMI[2].PAR.DRIVE.DIV_POS_SLOW := 60;
   HMI[2].PAR.DRIVE.TOL_SET_POS := 2;
   HMI[2].PAR.DRIVE.TOL_RESET_POS := 20;
   HMI[2].PAR.DRIVE.Window_Pos := 2;
   HMI[2].PAR.DRIVE.Window_Overrun := 10;
   HMI[2].PAR.DRIVE.Window_Pos_2 := 800;
   HMI[2].PAR.DRIVE.Window_Movement := 10;
   HMI[2].PAR.DRIVE.Window_Distance_Reserve := 10;
   HMI[2].PAR.DRIVE.Delay_Pos := 2000;
   HMI[2].PAR.DRIVE.Reserve_118 := S5T#5M;
   HMI[2].PAR.DRIVE.Reserve_120 := S5T#2M;
   HMI[2].PAR.DRIVE.DelaySpeedContr := S5T#6S_600MS;
   HMI[2].PAR.DRIVE.TolSpeedContr := 30;
   HMI[2].PAR.DRIVE.SYNCH_MID_VALUE := 0;
   HMI[2].PAR.Reserve[1] := 16#0000;
   HMI[2].PAR.Reserve[2] := 16#0000;
   HMI[2].PAR.Reserve[3] := 16#0000;
   HMI[2].PAR.Reserve[4] := 16#0000;
   HMI[2].PAR.Reserve[5] := 16#0000;
   HMI[2].PAR.HOIST.V_Min := 0;
   HMI[2].PAR.HOIST.V_Max := 8000;
   HMI[2].PAR.HOIST.V_MaxOccLift := 6500;
   HMI[2].PAR.HOIST.V_Reserve_2 := 0;
   HMI[2].PAR.HOIST.V_Pos_1 := 800;
   HMI[2].PAR.HOIST.V_Pos_2 := 2000;
   HMI[2].PAR.HOIST.V_Fixed_1 := 2000;
   HMI[2].PAR.HOIST.V_Fixed_2 := 4000;
   HMI[2].PAR.HOIST.V_Fixed_3_START := 400;
   // 2060 more start values not shown
END_DATA_BLOCK

DATA_BLOCK "DB_SDC_TS_PARAMETER_HMI"   // DB3804
{ S7_Optimized_Access := 'FALSE' }
AUTHOR : FFM
FAMILY : SDC
NAME : SECT_DEF
VERSION : 1.0
   VAR
      HEADER : Struct
         DB_NR : Int := 3804;
         Res020 : Int := 0;
         Res040 : Int := 0;
         START_DAT : Int := 20;
         LAENGE_SEK_DATA : Int := 480;
         ANZ_PROFIL : Int := 10;
         OFFEST_PROFIL : Int := 40;
         LAENGE_PROFIL_DATA : Int := 44;
         START_HMI : Int := 20;
         OFFEST_HMI_DATA : Int := 20;
      END_STRUCT;
      HMI : Array[1..30] of Struct
         PULT_Nr_EDIT : Int;
         BILD_Nr : Int;
         BILD_Nr_Alt : Int;
         SEK_Nr : Int;
         SEK_Nr_Alt : Int;
         PROFIL_Nr : Int;
         PROFIL_Nr_Alt : Int;
         PROFIL_Nr_COPY : Int;
         PROFIL_Nr_DEST : Int;
         T_EDIT : Bool;
         T_RESET_BED : Bool;
         T_SAVE : Bool;
         T_LOAD : Bool;
         T_COPY : Bool;
         T_COPY_ALL : Bool;
         Res086 : Bool;
         Res087 : Bool;
         FR_EDIT : Bool;
         ER_DATA : Bool;
         TS : "UDT_SDC_TS_PARAMETER";
      END_STRUCT;
   END_VAR
BEGIN
   HMI[19].PROFIL_Nr_COPY := 1;
   HMI[19].PROFIL_Nr_DEST := 2;
   HMI[18].PROFIL_Nr_COPY := 0;
   HMI[18].PROFIL_Nr_DEST := 0;
   HMI[1].PULT_Nr_EDIT := 0;
   HMI[1].BILD_Nr := 0;
   HMI[1].BILD_Nr_Alt := 0;
   HMI[1].SEK_Nr := 255;
   HMI[1].SEK_Nr_Alt := 255;
   HMI[1].PROFIL_Nr := 1;
   HMI[1].PROFIL_Nr_Alt := 1;
   HMI[1].PROFIL_Nr_COPY := 0;
   HMI[1].PROFIL_Nr_DEST := 0;
   HMI[1].T_EDIT := FALSE;
   HMI[1].T_RESET_BED := FALSE;
   HMI[1].T_SAVE := FALSE;
   HMI[1].T_LOAD := FALSE;
   HMI[1].T_COPY := FALSE;
   HMI[1].T_COPY_ALL := FALSE;
   HMI[1].Res086 := FALSE;
   HMI[1].Res087 := FALSE;
   HMI[1].FR_EDIT := FALSE;
   HMI[1].ER_DATA := FALSE;
   HMI[1].TS.ALLG.SEK_NEXT_1 := 0;
   HMI[1].TS.ALLG.SEK_NEXT_2 := 0;
   HMI[1].TS.ALLG.Spare[4] := 16#00;
   HMI[1].TS.ALLG.Spare[5] := 16#00;
   HMI[1].TS.ALLG.POS.Start_1 := 24601;
   HMI[1].TS.ALLG.POS.End_1 := 30800;
   HMI[1].TS.ALLG.POS.Start_2 := 0;
   HMI[1].TS.ALLG.POS.End_2 := 0;
   HMI[1].TS.ALLG.POS.Actionpoint_1 := 0;
   HMI[1].TS.ALLG.POS.Actionpoint_2 := 0;
   HMI[1].TS.ALLG.FLAGS.DIST_VAL[0] := TRUE;
   HMI[1].TS.ALLG.FLAGS.DIST_VAL[1] := FALSE;
   HMI[1].TS.ALLG.FLAGS.DIST_VAL[2] := FALSE;
   HMI[1].TS.ALLG.FLAGS.DIST_VAL[3] := FALSE;
   HMI[1].TS.ALLG.FLAGS.DIST_VAL[4] := FALSE;
   HMI[1].TS.ALLG.FLAGS.DIST_VAL[5] := FALSE;
   HMI[1].TS.ALLG.FLAGS.DIST_VAL[6] := FALSE;
   HMI[1].TS.ALLG.FLAGS.DIST_VAL[7] := FALSE;
   HMI[1].TS.ALLG.FLAGS.DIST_VAL[8] := FALSE;
   HMI[1].TS.ALLG.FLAGS.DIST_VAL[9] := FALSE;
   HMI[1].TS.ALLG.FLAGS.DIST_VAL[10] := FALSE;
   HMI[1].TS.ALLG.FLAGS.DIST_VAL[11] := FALSE;
   HMI[1].TS.ALLG.FLAGS.DIST_VAL[12] := FALSE;
   HMI[1].TS.ALLG.FLAGS.DIST_VAL[13] := FALSE;
   HMI[1].TS.ALLG.FLAGS.DIST_VAL[14] := FALSE;
   HMI[1].TS.ALLG.FLAGS.DIST_VAL[15] := FALSE;
   HMI[1].TS.ALLG.FLAGS.one_profile := FALSE;
   HMI[1].TS.ALLG.FLAGS.BLIND := FALSE;
   HMI[1].TS.ALLG.FLAGS.NO_DIST_CONT := FALSE;
   HMI[1].TS.ALLG.FLAGS.SYNCH_AREA := FALSE;
   HMI[1].TS.ALLG.FLAGS.bit24 := FALSE;
   HMI[1].TS.ALLG.FLAGS.bit25 := FALSE;
   HMI[1].TS.ALLG.FLAGS.bit26 := FALSE;
   HMI[1].TS.ALLG.FLAGS.bit27 := FALSE;
   HMI[1].TS.ALLG.FLAGS.EN_HOIST := TRUE;
   HMI[1].TS.ALLG.FLAGS.D_RESET_AFTER := FALSE;
   HMI[1].TS.ALLG.FLAGS.D_PULK := FALSE;
   HMI[1].TS.ALLG.FLAGS.bit33 := FALSE;
   HMI[1].TS.ALLG.FLAGS.bit34 := FALSE;
   HMI[1].TS.ALLG.FLAGS.bit35 := FALSE;
   HMI[1].TS.ALLG.FLAGS.bit36 := FALSE;
   HMI[1].TS.ALLG.FLAGS.Deutronic_ON := FALSE;
   HMI[1].TS.ALLG.Stop_Position := 3221;
   HMI[1].TS.ALLG.Drive_speed_1 := 16000;
   HMI[1].TS.ALLG.Drive_speed_2 := 16000;
   HMI[1].TS.PROFIL[1].Hoist_Pos_start := 0;
   HMI[1].TS.PROFIL[1].Height := 2747;
   HMI[1].TS.PROFIL[1].Hoist_speed := 0;
   HMI[1].TS.PROFIL[1].Hoist_offset_1 := 0;
   HMI[1].TS.PROFIL[1].Hoist_offset_2 := 0;
   HMI[1].TS.PROFIL[1].Hoist_offset_3 := 0;
   HMI[1].TS.PROFIL[1].Hoist_offset_4 := 0;
   HMI[1].TS.PROFIL[1].Hoist_Start_offset_1 := 0;
   HMI[1].TS.PROFIL[1].Hoist_Start_offset_2 := 0;
   HMI[1].TS.PROFIL[1].Hoist_Start_offset_3 := 0;
   HMI[1].TS.PROFIL[1].Hoist_Start_offset_4 := 0;
   HMI[1].TS.PROFIL[2].Hoist_Pos_start := 0;
   HMI[1].TS.PROFIL[2].Height := 2747;
   HMI[1].TS.PROFIL[2].Hoist_speed := 0;
   HMI[1].TS.PROFIL[2].Hoist_offset_1 := 0;
   HMI[1].TS.PROFIL[2].Hoist_offset_2 := 0;
   HMI[1].TS.PROFIL[2].Hoist_offset_3 := 0;
   HMI[1].TS.PROFIL[2].Hoist_offset_4 := 0;
   HMI[1].TS.PROFIL[2].Hoist_Start_offset_1 := 0;
   HMI[1].TS.PROFIL[2].Hoist_Start_offset_2 := 0;
   HMI[1].TS.PROFIL[2].Hoist_Start_offset_3 := 0;
   HMI[1].TS.PROFIL[2].Hoist_Start_offset_4 := 0;
   HMI[1].TS.PROFIL[3].Hoist_Pos_start := 0;
   HMI[1].TS.PROFIL[3].Height := 3113;
   HMI[1].TS.PROFIL[3].Hoist_speed := 0;
   HMI[1].TS.PROFIL[3].Hoist_offset_1 := 0;
   HMI[1].TS.PROFIL[3].Hoist_offset_2 := 0;
   HMI[1].TS.PROFIL[3].Hoist_offset_3 := 0;
   HMI[1].TS.PROFIL[3].Hoist_offset_4 := 0;
   HMI[1].TS.PROFIL[3].Hoist_Start_offset_1 := 0;
   HMI[1].TS.PROFIL[3].Hoist_Start_offset_2 := 0;
   HMI[1].TS.PROFIL[3].Hoist_Start_offset_3 := 0;
   HMI[1].TS.PROFIL[3].Hoist_Start_offset_4 := 0;
   HMI[1].TS.PROFIL[4].Hoist_Pos_start := 0;
   HMI[1].TS.PROFIL[4].Height := 3113;
   HMI[1].TS.PROFIL[4].Hoist_speed := 0;
   HMI[1].TS.PROFIL[4].Hoist_offset_1 := 0;
   HMI[1].TS.PROFIL[4].Hoist_offset_2 := 0;
   HMI[1].TS.PROFIL[4].Hoist_offset_3 := 0;
   HMI[1].TS.PROFIL[4].Hoist_offset_4 := 0;
   HMI[1].TS.PROFIL[4].Hoist_Start_offset_1 := 0;
   HMI[1].TS.PROFIL[4].Hoist_Start_offset_2 := 0;
   HMI[1].TS.PROFIL[4].Hoist_Start_offset_3 := 0;
   HMI[1].TS.PROFIL[4].Hoist_Start_offset_4 := 0;
   HMI[1].TS.PROFIL[5].Hoist_Pos_start := 0;
   HMI[1].TS.PROFIL[5].Height := 3113;
   HMI[1].TS.PROFIL[5].Hoist_speed := 0;
   HMI[1].TS.PROFIL[5].Hoist_offset_1 := 0;
   HMI[1].TS.PROFIL[5].Hoist_offset_2 := 0;
   HMI[1].TS.PROFIL[5].Hoist_offset_3 := 0;
   HMI[1].TS.PROFIL[5].Hoist_offset_4 := 0;
   HMI[1].TS.PROFIL[5].Hoist_Start_offset_1 := 0;
   HMI[1].TS.PROFIL[5].Hoist_Start_offset_2 := 0;
   HMI[1].TS.PROFIL[5].Hoist_Start_offset_3 := 0;
   HMI[1].TS.PROFIL[5].Hoist_Start_offset_4 := 0;
   HMI[1].TS.PROFIL[6].Hoist_Pos_start := 0;
   HMI[1].TS.PROFIL[6].Height := 3113;
   HMI[1].TS.PROFIL[6].Hoist_speed := 0;
   HMI[1].TS.PROFIL[6].Hoist_offset_1 := 0;
   HMI[1].TS.PROFIL[6].Hoist_offset_2 := 0;
   HMI[1].TS.PROFIL[6].Hoist_offset_3 := 0;
   HMI[1].TS.PROFIL[6].Hoist_offset_4 := 0;
   HMI[1].TS.PROFIL[6].Hoist_Start_offset_1 := 0;
   HMI[1].TS.PROFIL[6].Hoist_Start_offset_2 := 0;
   HMI[1].TS.PROFIL[6].Hoist_Start_offset_3 := 0;
   HMI[1].TS.PROFIL[6].Hoist_Start_offset_4 := 0;
   HMI[1].TS.PROFIL[7].Hoist_Pos_start := 0;
   HMI[1].TS.PROFIL[7].Height := 3113;
   HMI[1].TS.PROFIL[7].Hoist_speed := 0;
   HMI[1].TS.PROFIL[7].Hoist_offset_1 := 0;
   HMI[1].TS.PROFIL[7].Hoist_offset_2 := 0;
   HMI[1].TS.PROFIL[7].Hoist_offset_3 := 0;
   HMI[1].TS.PROFIL[7].Hoist_offset_4 := 0;
   HMI[1].TS.PROFIL[7].Hoist_Start_offset_1 := 0;
   HMI[1].TS.PROFIL[7].Hoist_Start_offset_2 := 0;
   HMI[1].TS.PROFIL[7].Hoist_Start_offset_3 := 0;
   HMI[1].TS.PROFIL[7].Hoist_Start_offset_4 := 0;
   HMI[1].TS.PROFIL[8].Hoist_Pos_start := 0;
   HMI[1].TS.PROFIL[8].Height := 3113;
   HMI[1].TS.PROFIL[8].Hoist_speed := 0;
   HMI[1].TS.PROFIL[8].Hoist_offset_1 := 0;
   HMI[1].TS.PROFIL[8].Hoist_offset_2 := 0;
   HMI[1].TS.PROFIL[8].Hoist_offset_3 := 0;
   HMI[1].TS.PROFIL[8].Hoist_offset_4 := 0;
   HMI[1].TS.PROFIL[8].Hoist_Start_offset_1 := 0;
   HMI[1].TS.PROFIL[8].Hoist_Start_offset_2 := 0;
   HMI[1].TS.PROFIL[8].Hoist_Start_offset_3 := 0;
   HMI[1].TS.PROFIL[8].Hoist_Start_offset_4 := 0;
   HMI[1].TS.PROFIL[9].Hoist_Pos_start := 0;
   HMI[1].TS.PROFIL[9].Height := 3113;
   HMI[1].TS.PROFIL[9].Hoist_speed := 0;
   HMI[1].TS.PROFIL[9].Hoist_offset_1 := 0;
   HMI[1].TS.PROFIL[9].Hoist_offset_2 := 0;
   HMI[1].TS.PROFIL[9].Hoist_offset_3 := 0;
   HMI[1].TS.PROFIL[9].Hoist_offset_4 := 0;
   HMI[1].TS.PROFIL[9].Hoist_Start_offset_1 := 0;
   HMI[1].TS.PROFIL[9].Hoist_Start_offset_2 := 0;
   HMI[1].TS.PROFIL[9].Hoist_Start_offset_3 := 0;
   HMI[1].TS.PROFIL[9].Hoist_Start_offset_4 := 0;
   HMI[1].TS.PROFIL[10].Hoist_Pos_start := 0;
   HMI[1].TS.PROFIL[10].Height := 3113;
   HMI[1].TS.PROFIL[10].Hoist_speed := 0;
   HMI[1].TS.PROFIL[10].Hoist_offset_1 := 0;
   HMI[1].TS.PROFIL[10].Hoist_offset_2 := 0;
   HMI[1].TS.PROFIL[10].Hoist_offset_3 := 0;
   HMI[1].TS.PROFIL[10].Hoist_offset_4 := 0;
   HMI[1].TS.PROFIL[10].Hoist_Start_offset_1 := 0;
   HMI[1].TS.PROFIL[10].Hoist_Start_offset_2 := 0;
   HMI[1].TS.PROFIL[10].Hoist_Start_offset_3 := 0;
   HMI[1].TS.PROFIL[10].Hoist_Start_offset_4 := 0;
   HMI[2].PULT_Nr_EDIT := 0;
   HMI[2].BILD_Nr := 0;
   HMI[2].BILD_Nr_Alt := 0;
   HMI[2].SEK_Nr := 260;
   HMI[2].SEK_Nr_Alt := 260;
   HMI[2].PROFIL_Nr := 1;
   HMI[2].PROFIL_Nr_Alt := 1;
   HMI[2].PROFIL_Nr_COPY := 9;
   HMI[2].PROFIL_Nr_DEST := 0;
   HMI[2].T_EDIT := FALSE;
   HMI[2].T_RESET_BED := FALSE;
   HMI[2].T_SAVE := FALSE;
   HMI[2].T_LOAD := FALSE;
   HMI[2].T_COPY := FALSE;
   HMI[2].T_COPY_ALL := FALSE;
   HMI[2].Res086 := FALSE;
   HMI[2].Res087 := FALSE;
   HMI[2].FR_EDIT := FALSE;
   HMI[2].ER_DATA := FALSE;
   HMI[2].TS.ALLG.SEK_NEXT_1 := 0;
   HMI[2].TS.ALLG.SEK_NEXT_2 := 0;
   HMI[2].TS.ALLG.Spare[4] := 16#00;
   // 3280 more start values not shown
END_DATA_BLOCK

DATA_BLOCK "DB_SDC_EMS_TS_1_HMI"   // DB3810
{ S7_Optimized_Access := 'FALSE' }
VERSION : 0.1
   VAR
      HEADER : Struct   // Struktur für Datenheader // nicht verschieben
         DB_NR : Int := 3810;   // DB Nummer
         MIN_NR_SEK : Int := 1;   // Niedrigste SEK Nummer im DB
         MAX_NR_SEK : Int := 200;   // Höchste SEK Nummer im DB
         START_DAT : Int := 20;   // Startadresse der SEK im DB
         LAENGE_EMS_SEK_STAT : Int := 34;   // Länge EMS Data
         ANZ_EMS_SEK_STAT : Int := 6;   // Anzahl EMS Data
         MIN_DIST_EMS : DInt := 6000;   // min Distance EMS
         Res16 : Int := 0;   // Reserve
         Res18 : Int := 0;   // Reserve
      END_STRUCT;
      SEK : Array[1..200] of "UDT_SDC_6EMS_TS_STAT_HMI";
   END_VAR
BEGIN
END_DATA_BLOCK

DATA_BLOCK "DB_SDC_EMS_TS_2_HMI"   // DB3811
{ S7_Optimized_Access := 'FALSE' }
VERSION : 0.1
   VAR
      HEADER : Struct   // Struktur für Datenheader // nicht verschieben
         DB_NR : Int := 3811;   // DB Nummer
         MIN_NR_SEK : Int := 201;   // Niedrigste SEK Nummer im DB
         MAX_NR_SEK : Int := 400;   // Höchste SEK Nummer im DB
         START_DAT : Int := 20;   // Startadresse der SEK im DB
         LAENGE_EMS_SEK_STAT : Int := 34;   // Länge EMS Data
         ANZ_EMS_SEK_STAT : Int := 6;   // Anzahl EMS Data
         MIN_DIST_EMS : DInt := 6000;   // min Distance EMS
         Res16 : Int := 0;   // Reserve
         Res18 : Int := 0;   // Reserve
      END_STRUCT;
      SEK : Array[201..400] of "UDT_SDC_6EMS_TS_STAT_HMI";
   END_VAR
BEGIN
END_DATA_BLOCK

